(* Logix 5000 project; controller TemplateV1R0 vendor 1 type 14 code 222 rev 33.11; software revision 33.00; part 4 of 5 *)
(* tags used below, declared in another part *)
   Alarm : AlarmGenerator[10];
   AlarmText : STRING[10];
(* UnitX_EMXXX, continued *)

ROUTINE _EP_12_Unholding   (* ladder *)
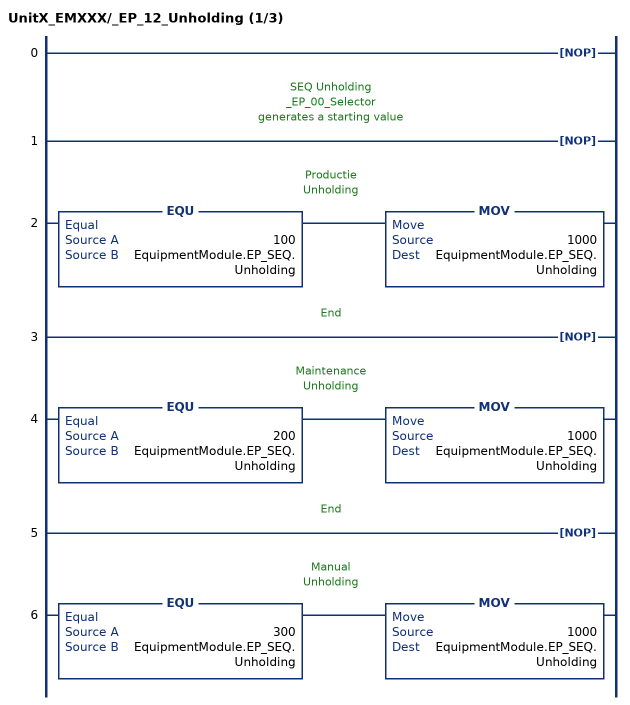
   0: NOP();
   // SEQ Unholding
   // _EP_00_Selector
   // generates a starting value
   1: NOP();
   // Productie
   // Unholding
   2: EQU(100,EquipmentModule.EP_SEQ.Unholding)MOV(1000,EquipmentModule.EP_SEQ.Unholding);
   // End
   3: NOP();
   // Maintenance
   // Unholding
   4: EQU(200,EquipmentModule.EP_SEQ.Unholding)MOV(1000,EquipmentModule.EP_SEQ.Unholding);
   // End
   5: NOP();
   // Manual
   // Unholding
   6: EQU(300,EquipmentModule.EP_SEQ.Unholding)MOV(1000,EquipmentModule.EP_SEQ.Unholding);
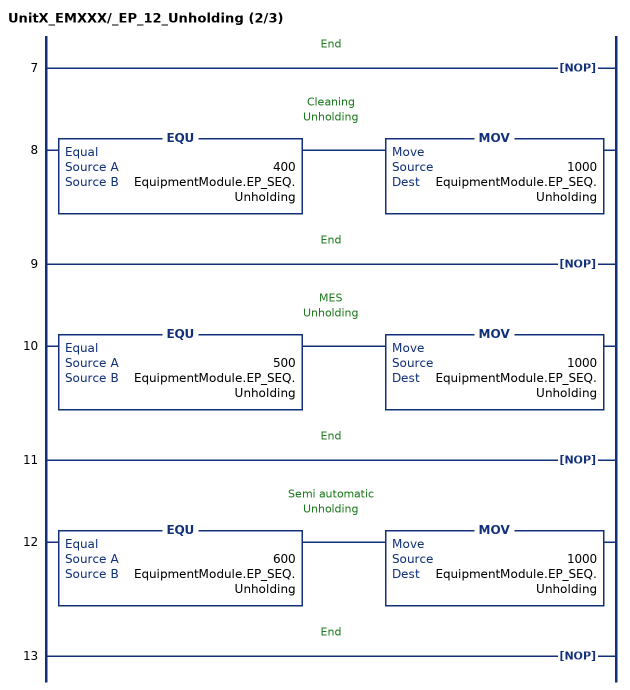
   // End
   7: NOP();
   // Cleaning
   // Unholding
   8: EQU(400,EquipmentModule.EP_SEQ.Unholding)MOV(1000,EquipmentModule.EP_SEQ.Unholding);
   // End
   9: NOP();
   // MES
   // Unholding
   10: EQU(500,EquipmentModule.EP_SEQ.Unholding)MOV(1000,EquipmentModule.EP_SEQ.Unholding);
   // End
   11: NOP();
   // Semi automatic
   // Unholding
   12: EQU(600,EquipmentModule.EP_SEQ.Unholding)MOV(1000,EquipmentModule.EP_SEQ.Unholding);
   // End
   13: NOP();
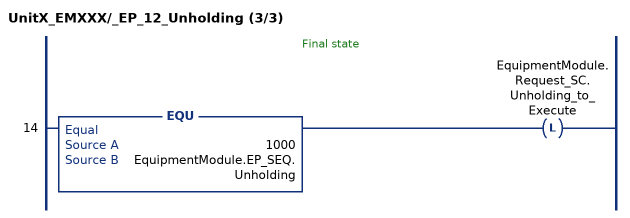
   // Final state
   14: EQU(1000,EquipmentModule.EP_SEQ.Unholding)OTL(EquipmentModule.Request_SC.Unholding_to_Execute);
END_ROUTINE

ROUTINE _EP_13_Suspending   (* ladder *)
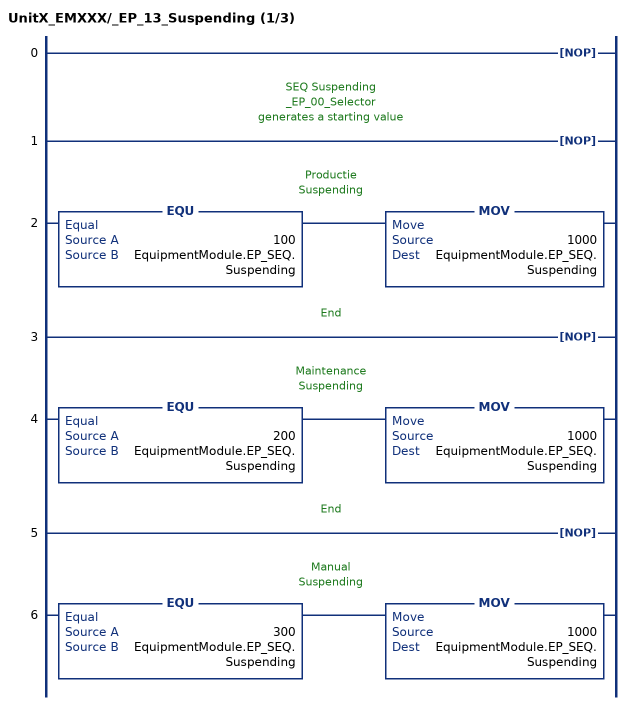
   0: NOP();
   // SEQ Suspending
   // _EP_00_Selector
   // generates a starting value
   1: NOP();
   // Productie
   // Suspending
   2: EQU(100,EquipmentModule.EP_SEQ.Suspending)MOV(1000,EquipmentModule.EP_SEQ.Suspending);
   // End
   3: NOP();
   // Maintenance
   // Suspending
   4: EQU(200,EquipmentModule.EP_SEQ.Suspending)MOV(1000,EquipmentModule.EP_SEQ.Suspending);
   // End
   5: NOP();
   // Manual
   // Suspending
   6: EQU(300,EquipmentModule.EP_SEQ.Suspending)MOV(1000,EquipmentModule.EP_SEQ.Suspending);
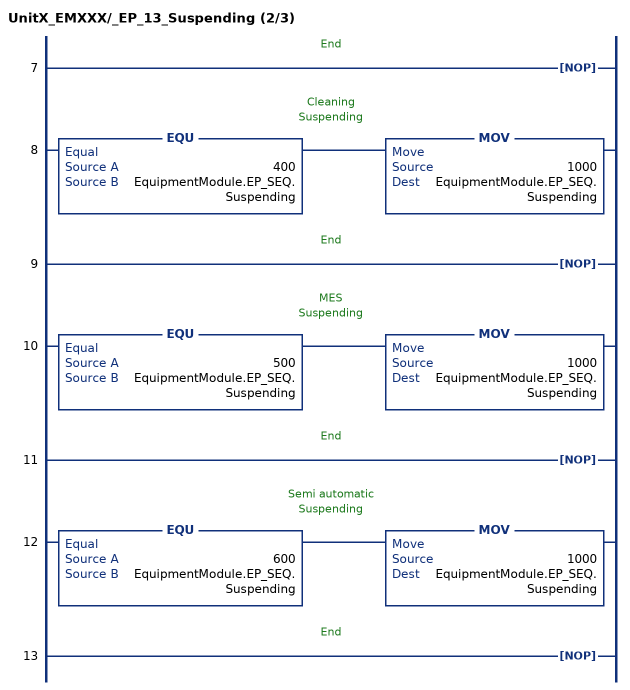
   // End
   7: NOP();
   // Cleaning
   // Suspending
   8: EQU(400,EquipmentModule.EP_SEQ.Suspending)MOV(1000,EquipmentModule.EP_SEQ.Suspending);
   // End
   9: NOP();
   // MES
   // Suspending
   10: EQU(500,EquipmentModule.EP_SEQ.Suspending)MOV(1000,EquipmentModule.EP_SEQ.Suspending);
   // End
   11: NOP();
   // Semi automatic
   // Suspending
   12: EQU(600,EquipmentModule.EP_SEQ.Suspending)MOV(1000,EquipmentModule.EP_SEQ.Suspending);
   // End
   13: NOP();
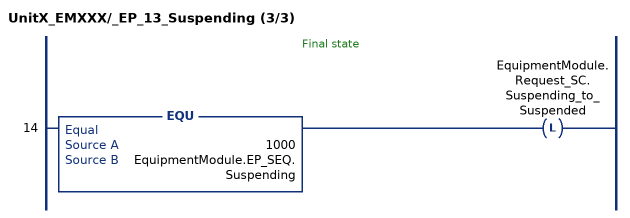
   // Final state
   14: EQU(1000,EquipmentModule.EP_SEQ.Suspending)OTL(EquipmentModule.Request_SC.Suspending_to_Suspended);
END_ROUTINE

ROUTINE _EP_14_Unsuspending   (* ladder *)
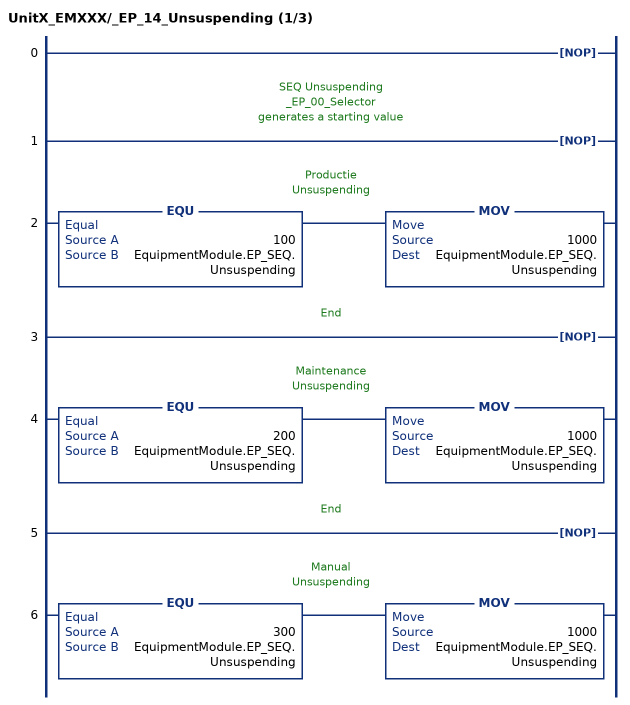
   0: NOP();
   // SEQ Unsuspending
   // _EP_00_Selector
   // generates a starting value
   1: NOP();
   // Productie
   // Unsuspending
   2: EQU(100,EquipmentModule.EP_SEQ.Unsuspending)MOV(1000,EquipmentModule.EP_SEQ.Unsuspending);
   // End
   3: NOP();
   // Maintenance
   // Unsuspending
   4: EQU(200,EquipmentModule.EP_SEQ.Unsuspending)MOV(1000,EquipmentModule.EP_SEQ.Unsuspending);
   // End
   5: NOP();
   // Manual
   // Unsuspending
   6: EQU(300,EquipmentModule.EP_SEQ.Unsuspending)MOV(1000,EquipmentModule.EP_SEQ.Unsuspending);
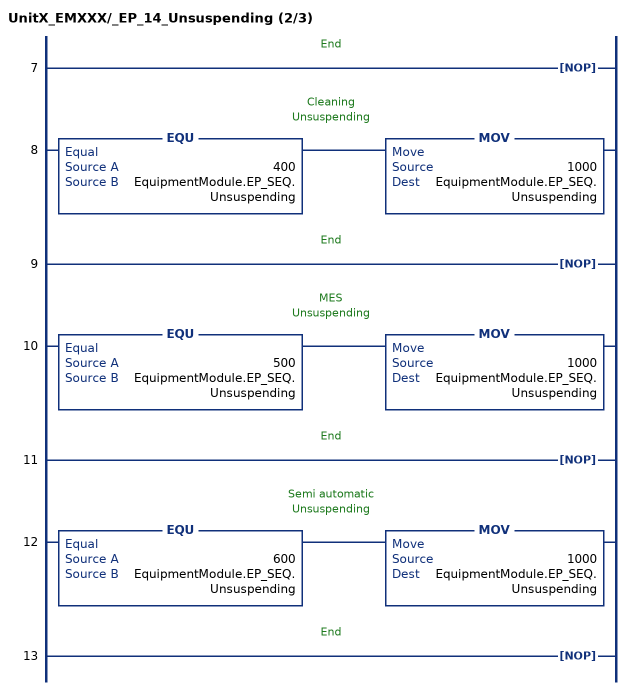
   // End
   7: NOP();
   // Cleaning
   // Unsuspending
   8: EQU(400,EquipmentModule.EP_SEQ.Unsuspending)MOV(1000,EquipmentModule.EP_SEQ.Unsuspending);
   // End
   9: NOP();
   // MES
   // Unsuspending
   10: EQU(500,EquipmentModule.EP_SEQ.Unsuspending)MOV(1000,EquipmentModule.EP_SEQ.Unsuspending);
   // End
   11: NOP();
   // Semi automatic
   // Unsuspending
   12: EQU(600,EquipmentModule.EP_SEQ.Unsuspending)MOV(1000,EquipmentModule.EP_SEQ.Unsuspending);
   // End
   13: NOP();
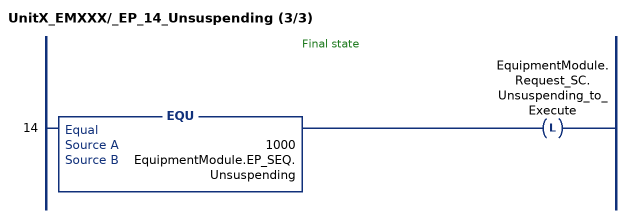
   // Final state
   14: EQU(1000,EquipmentModule.EP_SEQ.Unsuspending)OTL(EquipmentModule.Request_SC.Unsuspending_to_Execute);
END_ROUTINE

ROUTINE _EP_15_Resetting   (* ladder *)
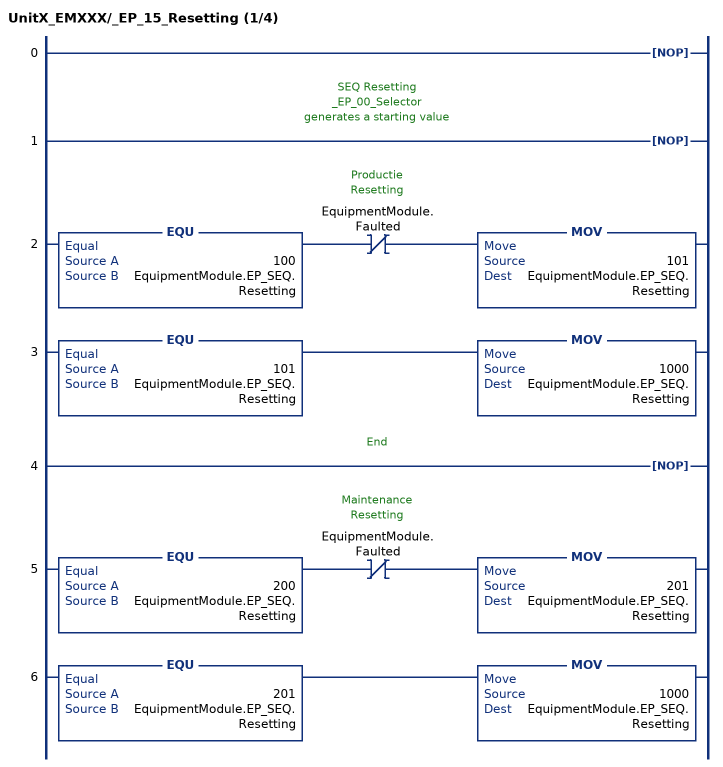
   0: NOP();
   // SEQ Resetting
   // _EP_00_Selector
   // generates a starting value
   1: NOP();
   // Productie
   // Resetting
   2: EQU(100,EquipmentModule.EP_SEQ.Resetting)XIO(EquipmentModule.Faulted)MOV(101,EquipmentModule.EP_SEQ.Resetting);
   3: EQU(101,EquipmentModule.EP_SEQ.Resetting)MOV(1000,EquipmentModule.EP_SEQ.Resetting);
   // End
   4: NOP();
   // Maintenance
   // Resetting
   5: EQU(200,EquipmentModule.EP_SEQ.Resetting)XIO(EquipmentModule.Faulted)MOV(201,EquipmentModule.EP_SEQ.Resetting);
   6: EQU(201,EquipmentModule.EP_SEQ.Resetting)MOV(1000,EquipmentModule.EP_SEQ.Resetting);
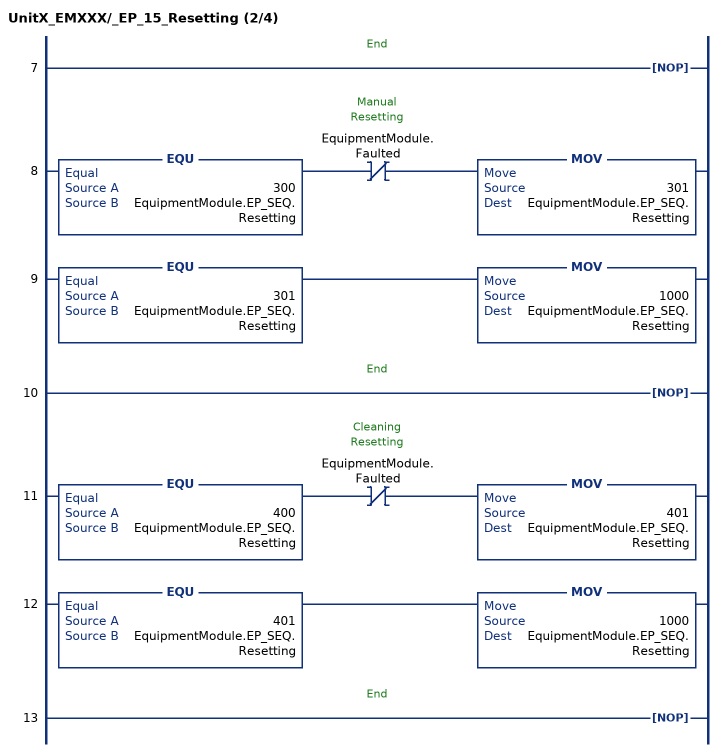
   // End
   7: NOP();
   // Manual
   // Resetting
   8: EQU(300,EquipmentModule.EP_SEQ.Resetting)XIO(EquipmentModule.Faulted)MOV(301,EquipmentModule.EP_SEQ.Resetting);
   9: EQU(301,EquipmentModule.EP_SEQ.Resetting)MOV(1000,EquipmentModule.EP_SEQ.Resetting);
   // End
   10: NOP();
   // Cleaning
   // Resetting
   11: EQU(400,EquipmentModule.EP_SEQ.Resetting)XIO(EquipmentModule.Faulted)MOV(401,EquipmentModule.EP_SEQ.Resetting);
   12: EQU(401,EquipmentModule.EP_SEQ.Resetting)MOV(1000,EquipmentModule.EP_SEQ.Resetting);
   // End
   13: NOP();
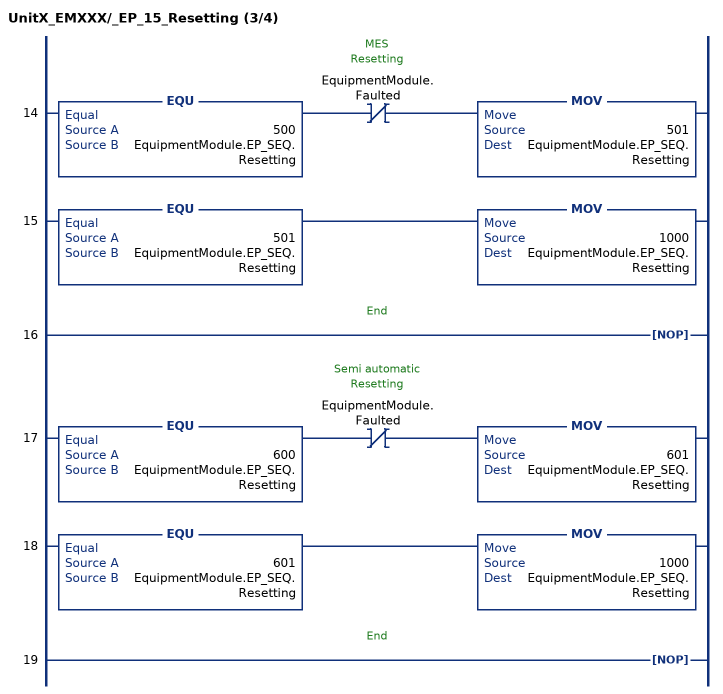
   // MES
   // Resetting
   14: EQU(500,EquipmentModule.EP_SEQ.Resetting)XIO(EquipmentModule.Faulted)MOV(501,EquipmentModule.EP_SEQ.Resetting);
   15: EQU(501,EquipmentModule.EP_SEQ.Resetting)MOV(1000,EquipmentModule.EP_SEQ.Resetting);
   // End
   16: NOP();
   // Semi automatic
   // Resetting
   17: EQU(600,EquipmentModule.EP_SEQ.Resetting)XIO(EquipmentModule.Faulted)MOV(601,EquipmentModule.EP_SEQ.Resetting);
   18: EQU(601,EquipmentModule.EP_SEQ.Resetting)MOV(1000,EquipmentModule.EP_SEQ.Resetting);
   // End
   19: NOP();
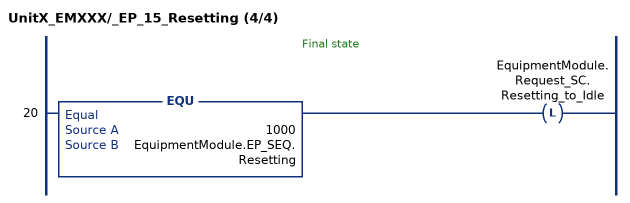
   // Final state
   20: EQU(1000,EquipmentModule.EP_SEQ.Resetting)OTL(EquipmentModule.Request_SC.Resetting_to_Idle);
END_ROUTINE

ROUTINE _EP_16_Completing   (* ladder *)
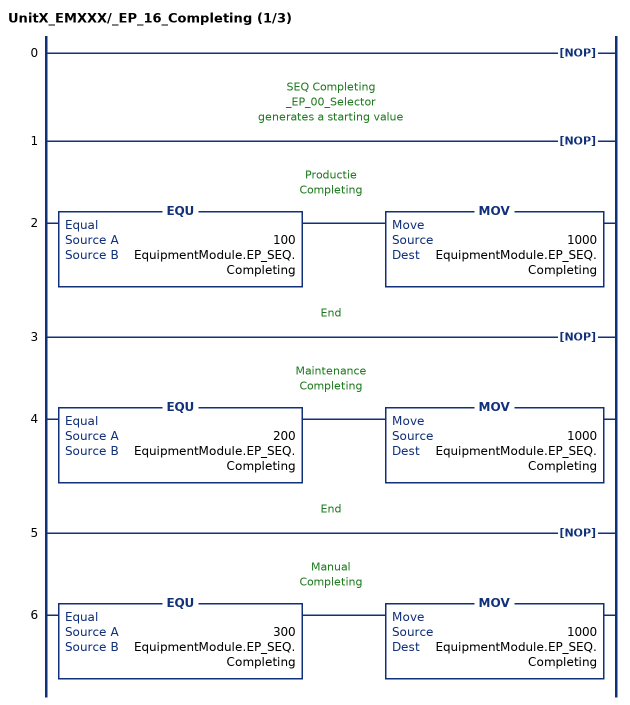
   0: NOP();
   // SEQ Completing
   // _EP_00_Selector
   // generates a starting value
   1: NOP();
   // Productie
   // Completing
   2: EQU(100,EquipmentModule.EP_SEQ.Completing)MOV(1000,EquipmentModule.EP_SEQ.Completing);
   // End
   3: NOP();
   // Maintenance
   // Completing
   4: EQU(200,EquipmentModule.EP_SEQ.Completing)MOV(1000,EquipmentModule.EP_SEQ.Completing);
   // End
   5: NOP();
   // Manual
   // Completing
   6: EQU(300,EquipmentModule.EP_SEQ.Completing)MOV(1000,EquipmentModule.EP_SEQ.Completing);
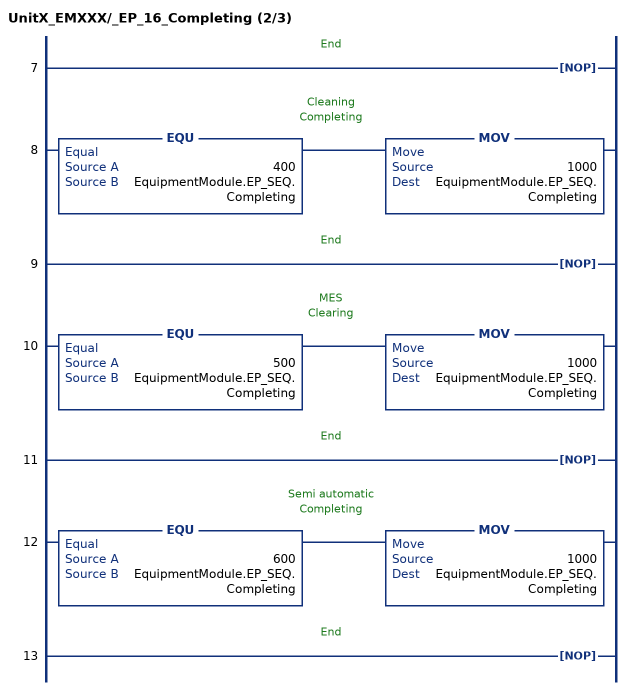
   // End
   7: NOP();
   // Cleaning
   // Completing
   8: EQU(400,EquipmentModule.EP_SEQ.Completing)MOV(1000,EquipmentModule.EP_SEQ.Completing);
   // End
   9: NOP();
   // MES
   // Clearing
   10: EQU(500,EquipmentModule.EP_SEQ.Completing)MOV(1000,EquipmentModule.EP_SEQ.Completing);
   // End
   11: NOP();
   // Semi automatic
   // Completing
   12: EQU(600,EquipmentModule.EP_SEQ.Completing)MOV(1000,EquipmentModule.EP_SEQ.Completing);
   // End
   13: NOP();
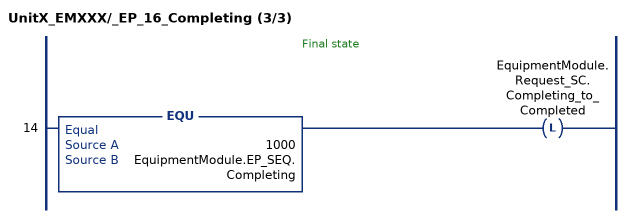
   // Final state
   14: EQU(1000,EquipmentModule.EP_SEQ.Completing)OTL(EquipmentModule.Request_SC.Completing_to_Completed);
END_ROUTINE

ROUTINE _FaultHandler   (* ladder *)
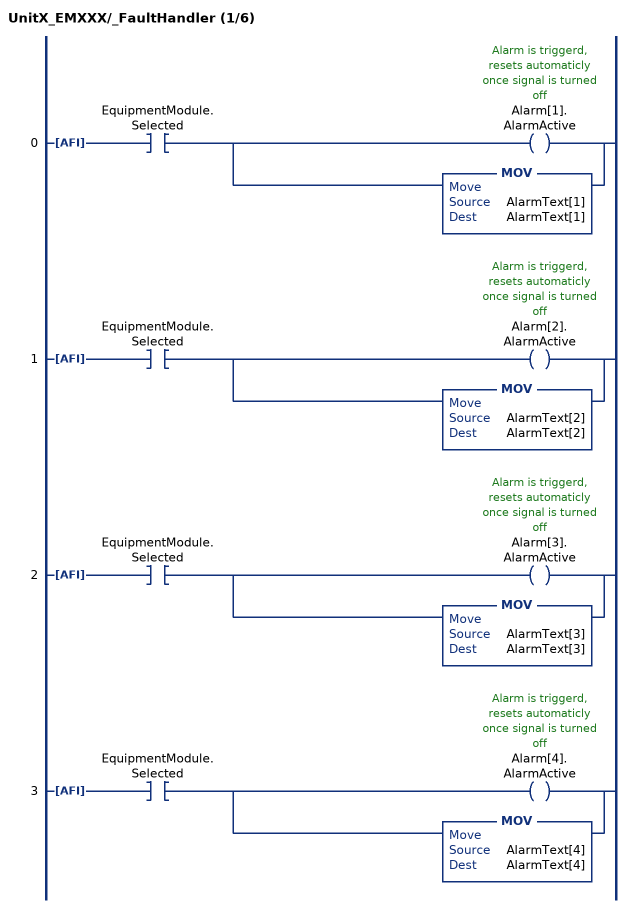
   0: AFI()XIC(EquipmentModule.Selected)[OTE(Alarm[1].AlarmActive) ,MOV(AlarmText[1],AlarmText[1]) ];
   1: AFI()XIC(EquipmentModule.Selected)[OTE(Alarm[2].AlarmActive) ,MOV(AlarmText[2],AlarmText[2]) ];
   2: AFI()XIC(EquipmentModule.Selected)[OTE(Alarm[3].AlarmActive) ,MOV(AlarmText[3],AlarmText[3]) ];
   3: AFI()XIC(EquipmentModule.Selected)[OTE(Alarm[4].AlarmActive) ,MOV(AlarmText[4],AlarmText[4]) ];
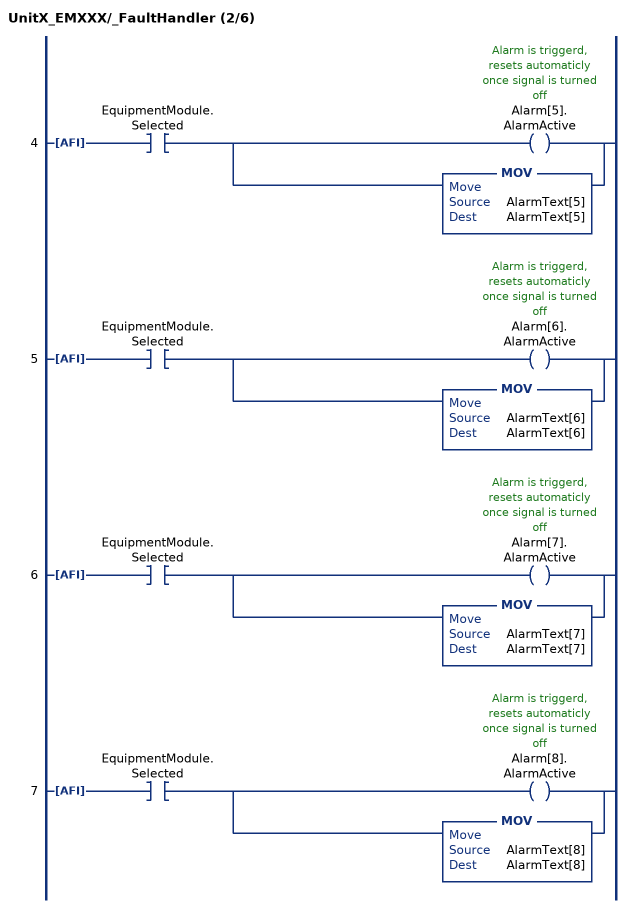
   4: AFI()XIC(EquipmentModule.Selected)[OTE(Alarm[5].AlarmActive) ,MOV(AlarmText[5],AlarmText[5]) ];
   5: AFI()XIC(EquipmentModule.Selected)[OTE(Alarm[6].AlarmActive) ,MOV(AlarmText[6],AlarmText[6]) ];
   6: AFI()XIC(EquipmentModule.Selected)[OTE(Alarm[7].AlarmActive) ,MOV(AlarmText[7],AlarmText[7]) ];
   7: AFI()XIC(EquipmentModule.Selected)[OTE(Alarm[8].AlarmActive) ,MOV(AlarmText[8],AlarmText[8]) ];
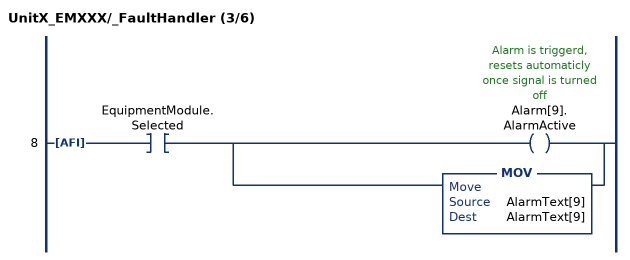
   8: AFI()XIC(EquipmentModule.Selected)[OTE(Alarm[9].AlarmActive) ,MOV(AlarmText[9],AlarmText[9]) ];
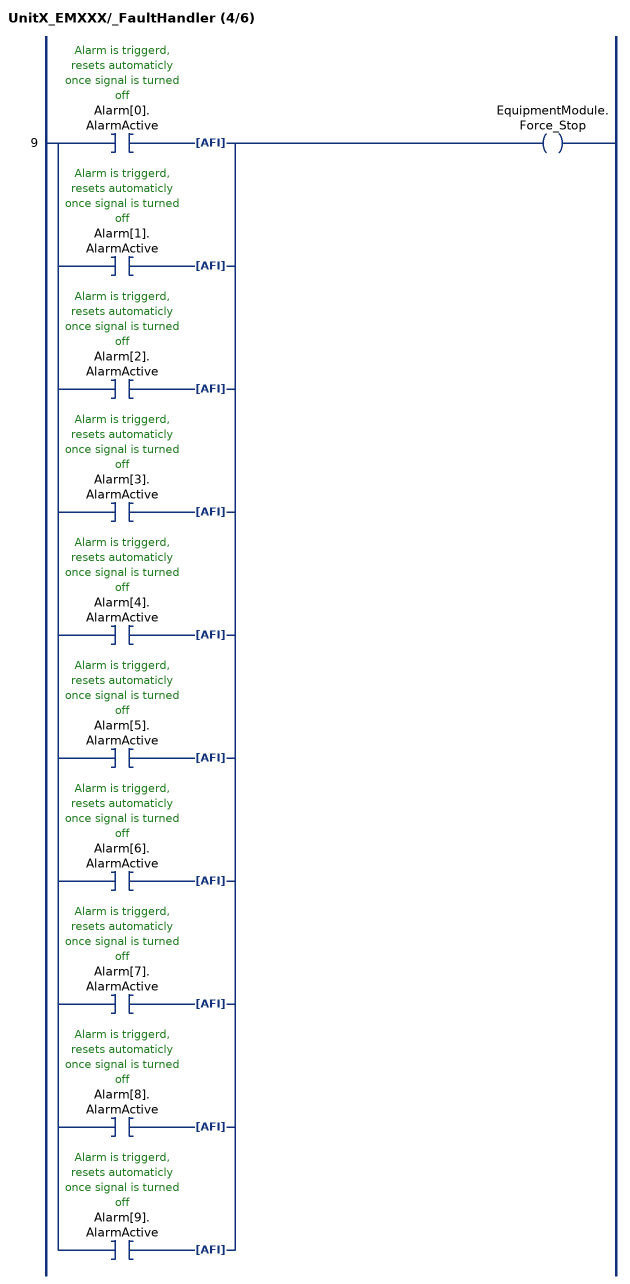
   9: [XIC(Alarm[0].AlarmActive) AFI() ,XIC(Alarm[1].AlarmActive) AFI() ,XIC(Alarm[2].AlarmActive) AFI() ,XIC(Alarm[3].AlarmActive) AFI() ,XIC(Alarm[4].AlarmActive) AFI() ,XIC(Alarm[5].AlarmActive) AFI() ,XIC(Alarm[6].AlarmActive) AFI() ,XIC(Alarm[7].AlarmActive) AFI() ,XIC(Alarm[8].AlarmActive) AFI() ,XIC(Alarm[9].AlarmActive) AFI() ]OTE(EquipmentModule.Force_Stop);
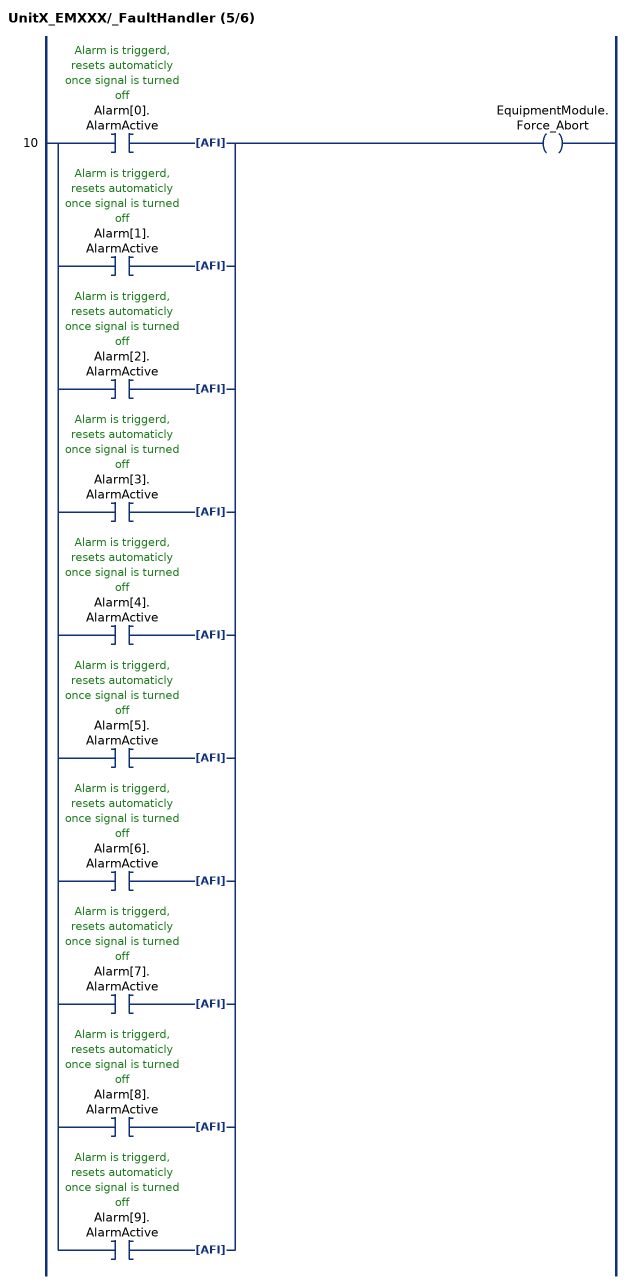
   10: [XIC(Alarm[0].AlarmActive) AFI() ,XIC(Alarm[1].AlarmActive) AFI() ,XIC(Alarm[2].AlarmActive) AFI() ,XIC(Alarm[3].AlarmActive) AFI() ,XIC(Alarm[4].AlarmActive) AFI() ,XIC(Alarm[5].AlarmActive) AFI() ,XIC(Alarm[6].AlarmActive) AFI() ,XIC(Alarm[7].AlarmActive) AFI() ,XIC(Alarm[8].AlarmActive) AFI() ,XIC(Alarm[9].AlarmActive) AFI() ]OTE(EquipmentModule.Force_Abort);
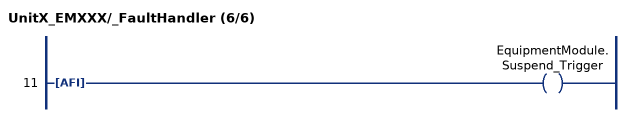
   11: AFI()OTE(EquipmentModule.Suspend_Trigger);
END_ROUTINE
